   END_RUNG
   RUNG wire#w1
      R_Coil( "PB Test Air Valve" )
   END_RUNG
   RUNG wire#w1
      R_Coil( "PB Test Pneumatic 6" )
   END_RUNG
   // the same network as SCL:
   #_w1 := NOT "Machine Running" AND NOT "PB Test Mode";
   IF #_w1 AND NOT "Error" THEN
       "Flag Yellow Light" := TRUE;
       "Flag Red Light" := FALSE;
       "Flag Green Light" := FALSE;
   END_IF;
   IF #_w1 AND NOT "Error" AND NOT "Error Door Open" AND NOT "Error Door Open FC" THEN
       "Flag Kran Angin" := TRUE;
   END_IF;
   IF #_w1 THEN
       "Flag Barcode Output" := FALSE;
       "Flag Pneumatic 1" := FALSE;
       "Flag Pneumatic 2" := FALSE;
       "Flag Pneumatic 3" := FALSE;
   END_IF;
   IF #_w1 AND NOT "Section Reject" THEN
       "Flag Pneumatic 4" := FALSE;
       "Flag Pneumatic 5" := FALSE;
   END_IF;
   IF #_w1 AND NOT "Slof Manual Ready" THEN "Flag Pneumatic 6" := FALSE; END_IF;
   IF #_w1 AND NOT "Section Reject" THEN "Flag Motor" := FALSE; END_IF;
   IF #_w1 THEN
       "Flag Imaje Start" := FALSE;
       "Flag Imaje Pause" := TRUE;
       "Flag Imaje Trigger" := FALSE;
       "Flag Mesin Sebelumnya" := FALSE;
       "PB Test Pneumatic 1" := FALSE;
       "PB Test Pneumatic 2" := FALSE;
       "PB Test Pneumatic 3" := FALSE;
       "PB Test Pneumatic 4" := FALSE;
       "PB Test Pneumatic 5" := FALSE;
       "PB Test Motor" := FALSE;
       "PB Test Imaje" := FALSE;
       "PB Test Air Valve" := FALSE;
       "PB Test Pneumatic 6" := FALSE;
   END_IF;
END_REGION

REGION Network 2: Output
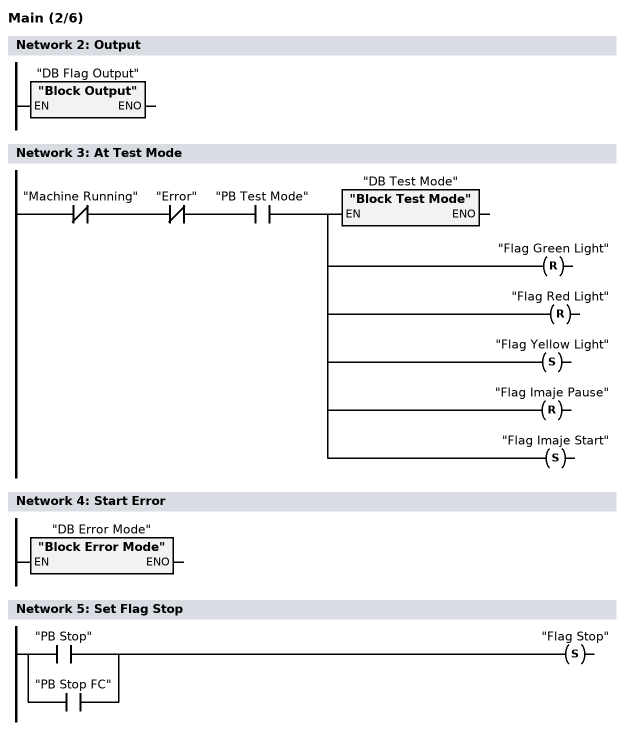
   RUNG wire#powerrail
      "DB Flag Output"()
   END_RUNG
   // the same network as SCL:
   "DB Flag Output"();   // "Block Output"
END_REGION

REGION Network 3: At Test Mode
   RUNG wire#powerrail
      I_Contact( "Machine Running" )
      I_Contact( "Error" )
      Contact( "PB Test Mode" )
      wire#w1
      "DB Test Mode"()
   END_RUNG
   RUNG wire#w1
      R_Coil( "Flag Green Light" )
   END_RUNG
   RUNG wire#w1
      R_Coil( "Flag Red Light" )
   END_RUNG
   RUNG wire#w1
      S_Coil( "Flag Yellow Light" )
   END_RUNG
   RUNG wire#w1
      R_Coil( "Flag Imaje Pause" )
   END_RUNG
   RUNG wire#w1
      S_Coil( "Flag Imaje Start" )
   END_RUNG
   // the same network as SCL:
   #_w1 := NOT "Machine Running" AND NOT "Error" AND "PB Test Mode";
   IF #_w1 THEN
       "DB Test Mode"();   // "Block Test Mode"
       "Flag Green Light" := FALSE;
       "Flag Red Light" := FALSE;
       "Flag Yellow Light" := TRUE;
       "Flag Imaje Pause" := FALSE;
       "Flag Imaje Start" := TRUE;
   END_IF;
END_REGION

REGION Network 4: Start Error
   RUNG wire#powerrail
      "DB Error Mode"()
   END_RUNG
   // the same network as SCL:
   "DB Error Mode"();   // "Block Error Mode"
END_REGION

REGION Network 5: Set Flag Stop
   RUNG wire#powerrail
      Contact( "PB Stop" )
      wire#w1
      S_Coil( "Flag Stop" )
   END_RUNG
   RUNG wire#powerrail
      Contact( "PB Stop FC" )
   END_RUNG wire#w1
   // the same network as SCL:
   IF "PB Stop" OR "PB Stop FC" THEN "Flag Stop" := TRUE; END_IF;
END_REGION

REGION Network 6: Flag Stop
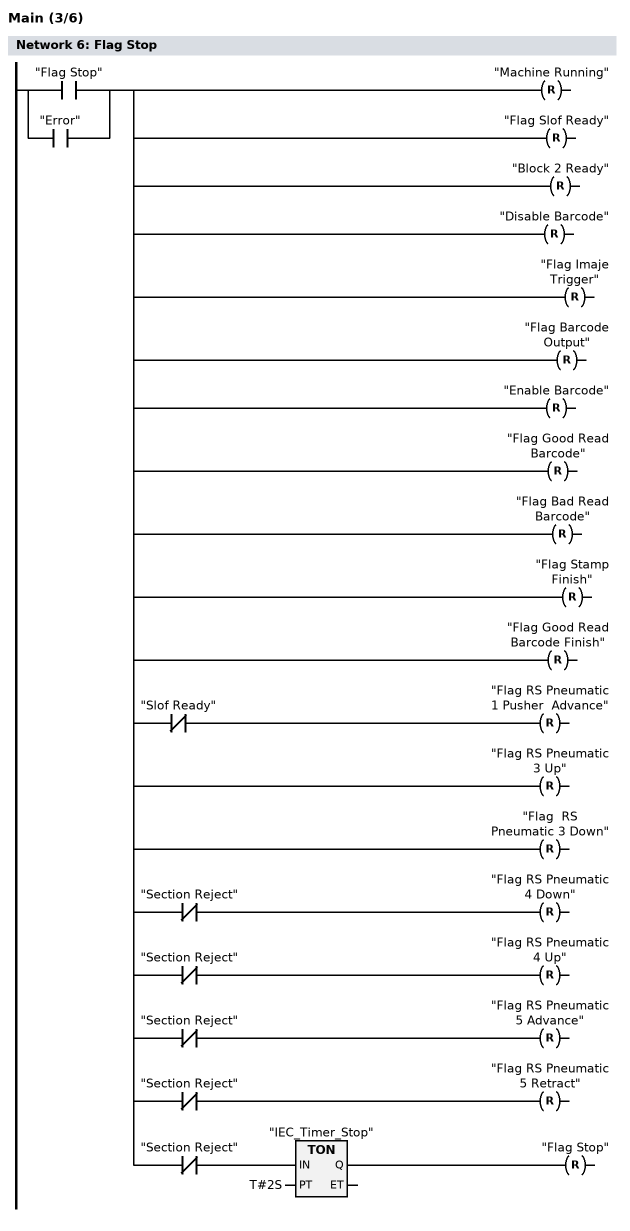
   #_w1 := "Flag Stop" OR "Error";
   IF #_w1 THEN
       "Machine Running" := FALSE;
       "Flag Slof Ready" := FALSE;
       "Block 2 Ready" := FALSE;
       "Disable Barcode" := FALSE;
       "Flag Imaje Trigger" := FALSE;
       "Flag Barcode Output" := FALSE;
       "Enable Barcode" := FALSE;
       "Flag Good Read Barcode" := FALSE;
       "Flag Bad Read Barcode" := FALSE;
       "Flag Stamp Finish" := FALSE;
       "Flag Good Read Barcode Finish" := FALSE;
   END_IF;
   IF #_w1 AND NOT "Slof Ready" THEN "Flag RS Pneumatic 1 Pusher  Advance" := FALSE; END_IF;
   IF #_w1 THEN
       "Flag RS Pneumatic 3 Up" := FALSE;
       "Flag  RS Pneumatic 3 Down" := FALSE;
   END_IF;
   IF #_w1 AND NOT "Section Reject" THEN
       "Flag RS Pneumatic 4 Down" := FALSE;
       "Flag RS Pneumatic 4 Up" := FALSE;
       "Flag RS Pneumatic 5 Advance" := FALSE;
       "Flag RS Pneumatic 5 Retract" := FALSE;
   END_IF;
   "IEC_Timer_Stop".TON(IN := #_w1 AND NOT "Section Reject", PT := T#2S);
   IF "IEC_Timer_Stop".Q THEN "Flag Stop" := FALSE; END_IF;
END_REGION

REGION Network 7: PB Run
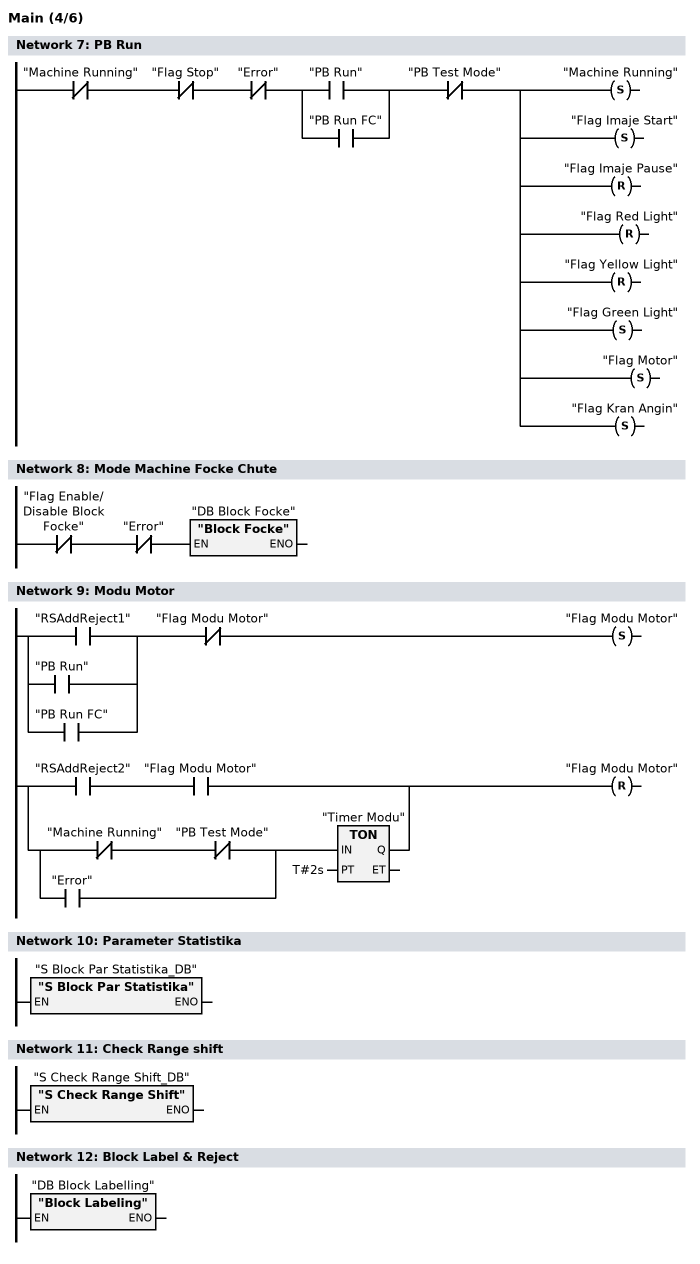
   RUNG wire#powerrail
      I_Contact( "Machine Running" )
      I_Contact( "Flag Stop" )
      I_Contact( "Error" )
      wire#w1
      Contact( "PB Run" )
      wire#w2
      I_Contact( "PB Test Mode" )
      wire#w3
      S_Coil( "Machine Running" )
   END_RUNG
   RUNG wire#w1
      Contact( "PB Run FC" )
   END_RUNG wire#w2
   RUNG wire#w3
      S_Coil( "Flag Imaje Start" )
   END_RUNG
   RUNG wire#w3
      R_Coil( "Flag Imaje Pause" )
   END_RUNG
   RUNG wire#w3
      R_Coil( "Flag Red Light" )
   END_RUNG
   RUNG wire#w3
      R_Coil( "Flag Yellow Light" )
   END_RUNG
   RUNG wire#w3
      S_Coil( "Flag Green Light" )
   END_RUNG
   RUNG wire#w3
      S_Coil( "Flag Motor" )
   END_RUNG
   RUNG wire#w3
      S_Coil( "Flag Kran Angin" )
   END_RUNG
   // the same network as SCL:
   #_w1 := NOT "Machine Running" AND NOT "Flag Stop" AND NOT "Error" AND ("PB Run" OR "PB Run FC") AND NOT "PB Test Mode";
   IF #_w1 THEN
       "Machine Running" := TRUE;
       "Flag Imaje Start" := TRUE;
       "Flag Imaje Pause" := FALSE;
       "Flag Red Light" := FALSE;
       "Flag Yellow Light" := FALSE;
       "Flag Green Light" := TRUE;
       "Flag Motor" := TRUE;
       "Flag Kran Angin" := TRUE;
   END_IF;
END_REGION

REGION Network 8: Mode Machine Focke Chute
   RUNG wire#powerrail
      I_Contact( "Flag Enable/Disable Block Focke" )
      I_Contact( "Error" )
      "DB Block Focke"()
   END_RUNG
   // the same network as SCL:
   IF NOT "Flag Enable/Disable Block Focke" AND NOT "Error" THEN
       "DB Block Focke"();   // "Block Focke"
   END_IF;
END_REGION

REGION Network 9: Modu Motor
   IF ("RSAddReject1" OR "PB Run" OR "PB Run FC") AND NOT "Flag Modu Motor" THEN
       "Flag Modu Motor" := TRUE;
   END_IF;
   "Timer Modu".TON(IN := (NOT "Machine Running" AND NOT "PB Test Mode") OR "Error", PT := T#2s);
   IF ("RSAddReject2" AND "Flag Modu Motor") OR "Timer Modu".Q THEN "Flag Modu Motor" := FALSE; END_IF;
END_REGION

REGION Network 10: Parameter Statistika
   RUNG wire#powerrail
      "S Block Par Statistika_DB"()
   END_RUNG
   // the same network as SCL:
   "S Block Par Statistika_DB"();   // "S Block Par Statistika"
END_REGION

REGION Network 11: Check Range shift
   RUNG wire#powerrail
      "S Check Range Shift_DB"()
   END_RUNG
   // the same network as SCL:
   "S Check Range Shift_DB"();   // "S Check Range Shift"
END_REGION

REGION Network 12: Block Label & Reject
   RUNG wire#powerrail
      "DB Block Labelling"()
   END_RUNG
   // the same network as SCL:
   "DB Block Labelling"();   // "Block Labeling"
END_REGION

REGION Network 13: Baca Data Statistika
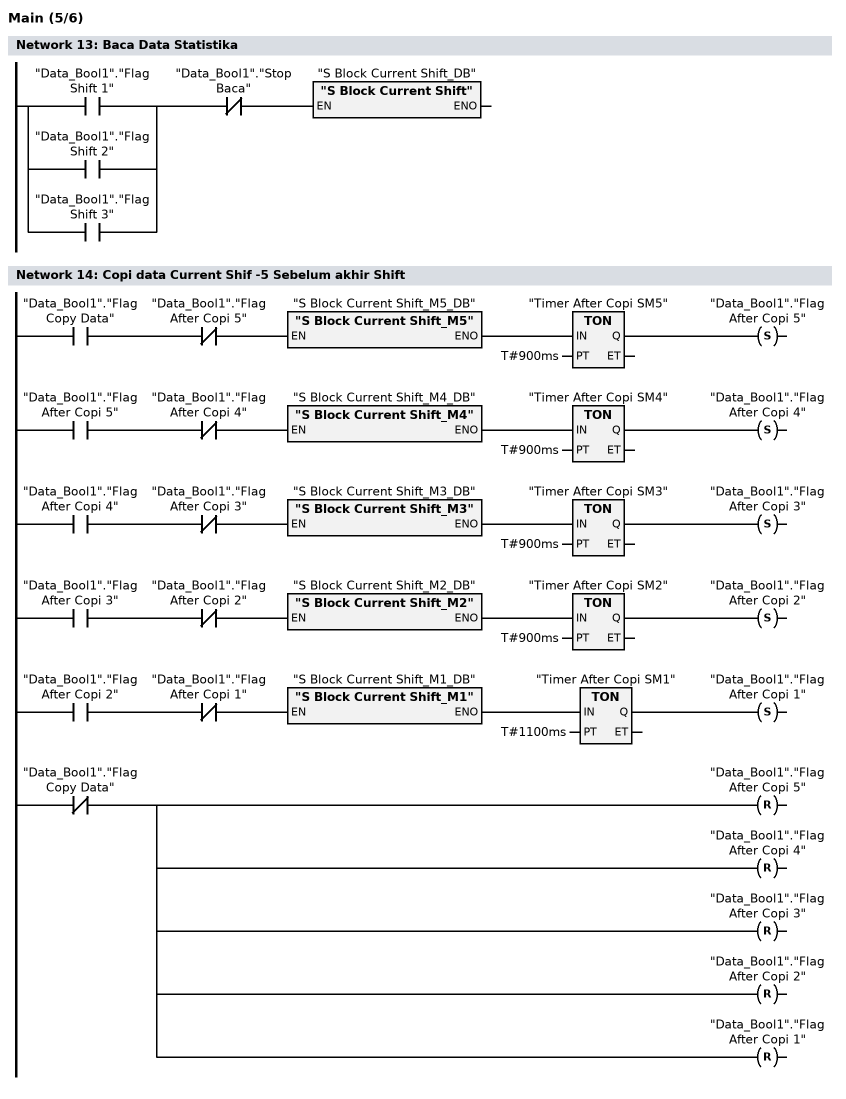
   RUNG wire#powerrail
      Contact( "Data_Bool1"."Flag Shift 1" )
      wire#w1
      I_Contact( "Data_Bool1"."Stop Baca" )
      "S Block Current Shift_DB"()
   END_RUNG
   RUNG wire#powerrail
      Contact( "Data_Bool1"."Flag Shift 2" )
   END_RUNG wire#w1
   RUNG wire#powerrail
      Contact( "Data_Bool1"."Flag Shift 3" )
   END_RUNG wire#w1
   // the same network as SCL:
   IF ("Data_Bool1"."Flag Shift 1" OR "Data_Bool1"."Flag Shift 2" OR "Data_Bool1"."Flag Shift 3") AND NOT "Data_Bool1"."Stop Baca" THEN
       "S Block Current Shift_DB"();   // "S Block Current Shift"
   END_IF;
END_REGION

REGION Network 14: Copi data Current Shif -5 Sebelum akhir Shift
   "S Block Current Shift_M5_DB"(EN := "Data_Bool1"."Flag Copy Data" AND NOT "Data_Bool1"."Flag After Copi 5",   // "S Block Current Shift_M5"
                           ENO => #_w1);
   "Timer After Copi SM5".TON(IN := #_w1, PT := T#900ms);
   IF "Timer After Copi SM5".Q THEN "Data_Bool1"."Flag After Copi 5" := TRUE; END_IF;
   "S Block Current Shift_M4_DB"(EN := "Data_Bool1"."Flag After Copi 5" AND NOT "Data_Bool1"."Flag After Copi 4",   // "S Block Current Shift_M4"
                           ENO => #_w2);
   "Timer After Copi SM4".TON(IN := #_w2, PT := T#900ms);
   IF "Timer After Copi SM4".Q THEN "Data_Bool1"."Flag After Copi 4" := TRUE; END_IF;
   "S Block Current Shift_M3_DB"(EN := "Data_Bool1"."Flag After Copi 4" AND NOT "Data_Bool1"."Flag After Copi 3",   // "S Block Current Shift_M3"
                           ENO => #_w3);
   "Timer After Copi SM3".TON(IN := #_w3, PT := T#900ms);
   IF "Timer After Copi SM3".Q THEN "Data_Bool1"."Flag After Copi 3" := TRUE; END_IF;
   "S Block Current Shift_M2_DB"(EN := "Data_Bool1"."Flag After Copi 3" AND NOT "Data_Bool1"."Flag After Copi 2",   // "S Block Current Shift_M2"
                           ENO => #_w4);
   "Timer After Copi SM2".TON(IN := #_w4, PT := T#900ms);
   IF "Timer After Copi SM2".Q THEN "Data_Bool1"."Flag After Copi 2" := TRUE; END_IF;
   "S Block Current Shift_M1_DB"(EN := "Data_Bool1"."Flag After Copi 2" AND NOT "Data_Bool1"."Flag After Copi 1",   // "S Block Current Shift_M1"
                           ENO => #_w5);
   "Timer After Copi SM1".TON(IN := #_w5, PT := T#1100ms);
   IF "Timer After Copi SM1".Q THEN "Data_Bool1"."Flag After Copi 1" := TRUE; END_IF;
   IF NOT "Data_Bool1"."Flag Copy Data" THEN
       "Data_Bool1"."Flag After Copi 5" := FALSE;
       "Data_Bool1"."Flag After Copi 4" := FALSE;
       "Data_Bool1"."Flag After Copi 3" := FALSE;
       "Data_Bool1"."Flag After Copi 2" := FALSE;
       "Data_Bool1"."Flag After Copi 1" := FALSE;
   END_IF;
END_REGION

REGION Network 15: Hapus Data Current shift
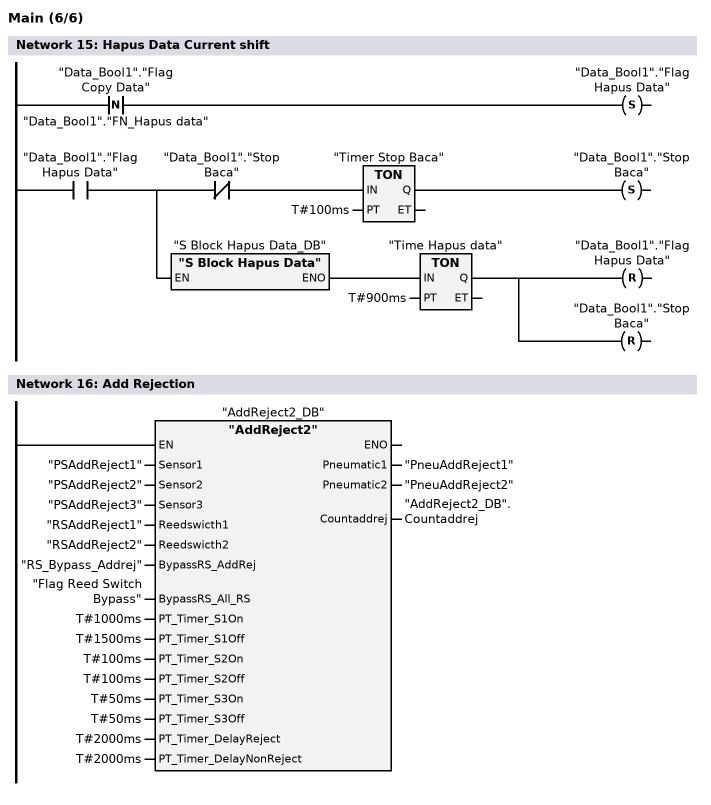
   #_w1 := NOT "Data_Bool1"."Flag Copy Data" AND "Data_Bool1"."FN_Hapus data";   // falling edge of "Data_Bool1"."Flag Copy Data"
   "Data_Bool1"."FN_Hapus data" := "Data_Bool1"."Flag Copy Data";
   IF #_w1 THEN "Data_Bool1"."Flag Hapus Data" := TRUE; END_IF;
   "Timer Stop Baca".TON(IN := "Data_Bool1"."Flag Hapus Data" AND NOT "Data_Bool1"."Stop Baca", PT := T#100ms);
   IF "Timer Stop Baca".Q THEN "Data_Bool1"."Stop Baca" := TRUE; END_IF;
   "S Block Hapus Data_DB"(EN := "Data_Bool1"."Flag Hapus Data", ENO => #_w2);   // "S Block Hapus Data"
   "Time Hapus data".TON(IN := #_w2, PT := T#900ms);
   IF "Time Hapus data".Q THEN
       "Data_Bool1"."Flag Hapus Data" := FALSE;
       "Data_Bool1"."Stop Baca" := FALSE;
   END_IF;
END_REGION

REGION Network 16: Add Rejection
   RUNG wire#powerrail
      "AddReject2_DB"(Sensor1 := "PSAddReject1", Sensor2 := "PSAddReject2", Sensor3 := "PSAddReject3", Reedswicth1 := "RSAddReject1", Reedswicth2 := "RSAddReject2", BypassRS_AddRej := "RS_Bypass_Addrej", BypassRS_All_RS := "Flag Reed Switch Bypass", PT_Timer_S1On := T#1000ms, PT_Timer_S1Off := T#1500ms, PT_Timer_S2On := T#100ms, PT_Timer_S2Off := T#100ms, PT_Timer_S3On := T#50ms, PT_Timer_S3Off := T#50ms, PT_Timer_DelayReject := T#2000ms, PT_Timer_DelayNonReject := T#2000ms, Pneumatic1 => "PneuAddReject1", Pneumatic2 => "PneuAddReject2", Countaddrej => "AddReject2_DB".Countaddrej)
   END_RUNG
   // the same network as SCL:
   "AddReject2_DB"(Sensor1 := "PSAddReject1",   // "AddReject2"
                   Sensor2 := "PSAddReject2",
                   Sensor3 := "PSAddReject3",
                   Reedswicth1 := "RSAddReject1",
                   Reedswicth2 := "RSAddReject2",
                   BypassRS_AddRej := "RS_Bypass_Addrej",
                   BypassRS_All_RS := "Flag Reed Switch Bypass",
                   PT_Timer_S1On := T#1000ms,
                   PT_Timer_S1Off := T#1500ms,
                   PT_Timer_S2On := T#100ms,
                   PT_Timer_S2Off := T#100ms,
                   PT_Timer_S3On := T#50ms,
                   PT_Timer_S3Off := T#50ms,
                   PT_Timer_DelayReject := T#2000ms,
                   PT_Timer_DelayNonReject := T#2000ms,
                   Pneumatic1 => "PneuAddReject1",
                   Pneumatic2 => "PneuAddReject2",
                   Countaddrej => "AddReject2_DB".Countaddrej);
END_REGION
END_ORGANIZATION_BLOCK

(* ===== HMI "HMI_RT_1" =====
system functions are stored by id; their names below are inferred from use
connection "HMI_connection": ETHERNET, SMART_S7_1200_OMS

HMI tags "Default tag table"
   "Tag_ScreenNumber" : UInt, internal
      on ChangeValue: ActivateScreenByNumber("Tag_ScreenNumber", 0)
   "PB Test Pneumatic 1" : Bool = PLC "PB Test Pneumatic 1" AT %M205.1, 1 s
   "PB Test Pneumatic 2" : Bool = PLC "PB Test Pneumatic 2" AT %M205.2, 1 s
   "PB Test Pneumatic 3" : Bool = PLC "PB Test Pneumatic 3" AT %M205.3, 1 s
   "PB Test Pneumatic 4" : Bool = PLC "PB Test Pneumatic 4" AT %M205.4, 1 s
   "PB Test Pneumatic 5" : Bool = PLC "PB Test Pneumatic 5" AT %M205.5, 1 s
   "PB Test Motor" : Bool = PLC "PB Test Motor" AT %M205.7, 1 s
   "PB Test Manual Servo" : Bool = PLC "PB Test Manual Servo" AT %M205.6, 1 s
   "Machine Running" : Bool = PLC "Machine Running" AT %M200.0, 1 s
   "Flag Imaje Start" : Bool = PLC "Flag Imaje Start" AT %M212.0, 1 s
   "Reset Counter" : Bool = PLC "Reset Counter" AT %M200.1, 1 s
   "PB Test Mode" : Bool = PLC "PB Test Mode" AT %M205.0, 1 s
   "Flag Ejector Jalan" : Bool = PLC "Flag Ejector Jalan" AT %M230.3, 1 s
   "Error Group" : Word = PLC "Error Group" AT %MW4, 1 s
   "PB Test Imaje" : Bool = PLC "PB Test Imaje" AT %M206.0, 1 s
   "PB Test Air Valve" : Bool = PLC "PB Test Air Valve" AT %M206.1, 1 s
   "Flag Barcode HMI" : Bool = PLC "Flag Enable/Disable Barcode HMI" AT %M30.0, 1 s
   "Flag Enable/Disable Error Chute 3 Way" : Bool = PLC "Flag Enable/Disable Error Chute 3 Way" AT %M30.1, 1 s
   "Flag Parameter Page" : Bool = PLC "Flag Parameter Page" AT %M232.6, 1 s
   "Flag Main Page" : Bool = PLC "Flag Main Page" AT %M232.7, 1 s
   "HMI_Tag_1" : Word AT %DB39.DBW0, 1 s
   "HMI_Error_Cont" : Word AT %DB40.DBW0, 1 s
   "Flag Teach In Barcode" : Bool = PLC "Flag Teach In Barcode" AT %M212.4, 1 s
   "Teach In Barcode" : Bool = PLC "Teach In Barcode" AT %Q0.5, 1 s
   "Flag Heater Error HMI" : Bool = PLC "Flag Heater Error HMI" AT %M30.2, 1 s
   "Flag Pneumatic Bypass" : Bool = PLC "Flag Reed Switch Bypass" AT %M30.3, 1 s
   "Flag Enable/Disable Error Door Open" : Bool = PLC "Flag Enable/Disable Error Door Open" AT %M30.5, 1 s
   "Flag Enable/Disable Block Focke" : Bool = PLC "Flag Enable/Disable Block Focke" AT %M30.6, 1 s
   "Flag Enable/Disable Error Chute Before Heating Roll" : Bool = PLC "Flag Enable/Disable Error Chute Before Heating Roll" AT %M30.4, 1 s
   "Flag Machine Bypass" : Bool = PLC "Flag Machine Bypass" AT %M30.7, 1 s
   "RS Bypass Pneumatic 1" : Bool = PLC "RS Bypass Pneumatic 1" AT %M31.0, 1 s
   "RS Bypass Pneumatic 3" : Bool = PLC "RS Bypass Pneumatic 3" AT %M31.1, 1 s
   "RS Bypass Pneumatic 4" : Bool = PLC "RS Bypass Pneumatic 4" AT %M31.2, 1 s
   "RS Bypass Pneumatic 5" : Bool = PLC "RS Bypass Pneumatic 5" AT %M31.3, 1 s
   "PB Test Pneumatic 6" : Bool = PLC "PB Test Pneumatic 6" AT %M206.2, 1 s
   "PB Test Conveyor" : Bool = PLC "PB Test Conveyor" AT %M206.3, 1 s
   "Flag Enable/Disable Flow to Reject" : Bool = PLC "Flag Enable/Disable Flow to Reject" AT %M31.5, 1 s
   "PB Test Motor Coveyor Pusher" : Bool = PLC "PB Test Motor Coveyor Pusher" AT %M206.4, 1 s
   "PB Test Motor Heating Roll" : Bool = PLC "PB Test Motor Heating Roll" AT %M206.5, 1 s
   "Flag Enable/Disable Heating Roll" : Bool = PLC "Flag Enable/Disable Heating Roll" AT %M31.6, 1 s
   "Flag Enable/Disable Reject Outfeed" : Bool = PLC "Flag Enable/Disable Reject Outfeed" AT %M31.7, 1 s
   "Data_DTL1_Output" : DTL = PLC Data_DTL1.Output, 1 s
   "Data_DTL1_Cur_ShiftA" : DTL = PLC Data_DTL1.Cur_ShiftA, 1 s
   "Data_DTL1_Cur_ShiftB" : DTL = PLC Data_DTL1.Cur_ShiftB, 1 s
   "Data_IntData_Input Sloft" : UDInt = PLC Data_IntData."Input Sloft", 1 s
   "Data_IntData_Tot Out Slof" : UDInt = PLC Data_IntData."Tot Out Slof", 1 s
   "Data_IntData_Good R" : UDInt = PLC Data_IntData."Good R", 1 s
   "Data_IntData_Reject Out S" : UDInt = PLC Data_IntData."Reject Out S", 1 s
   "Data_IntData_Bad R" : UDInt = PLC Data_IntData."Bad R", 1 s
   "Data_Real_% Total Output[0]" : Real = PLC Data_Real."% Total Output"[0], 1 s
   "Data_Real_%Good Read[0]" : Real = PLC Data_Real."%Good Read"[0], 1 s
   "Data_Real_% Reject Out Stop[0]" : Real = PLC Data_Real."% Reject Out Stop"[0], 1 s
   "Data_Real_%Bad Read[0]" : Real = PLC Data_Real."%Bad Read"[0], 1 s
   "Data_DTL1_Cur_ShiftA_1" : DTL = PLC Data_DTL1.Cur_ShiftA_1, 1 s
   "Data_DTL1_Cur_ShiftB_1" : DTL = PLC Data_DTL1.Cur_ShiftB_1, 1 s
   "Data_DTL1_Cur_ShiftA_2" : DTL = PLC Data_DTL1.Cur_ShiftA_2, 1 s
   "Data_DTL1_Cur_ShiftB_2" : DTL = PLC Data_DTL1.Cur_ShiftB_2, 1 s
   "Data_DTL1_Cur_ShiftA_3" : DTL = PLC Data_DTL1.Cur_ShiftA_3, 1 s
   "Data_DTL1_Cur_ShiftB_3" : DTL = PLC Data_DTL1.Cur_ShiftB_3, 1 s
   "Data_DTL1_Cur_ShiftA_4" : DTL = PLC Data_DTL1.Cur_ShiftA_4, 1 s
   "Data_DTL1_Cur_ShiftB_4" : DTL = PLC Data_DTL1.Cur_ShiftB_4, 1 s
   "Data_IntData_Input Sloft_1" : UDInt = PLC Data_IntData."Input Sloft_1", 1 s
   "Data_IntData_Tot Out Slof_1" : UDInt = PLC Data_IntData."Tot Out Slof_1", 1 s
   "Data_IntData_Good R_1" : UDInt = PLC Data_IntData."Good R_1", 1 s
   "Data_IntData_Reject Out S_1" : UDInt = PLC Data_IntData."Reject Out S_1", 1 s
   "Data_IntData_Bad R_1" : UDInt = PLC Data_IntData."Bad R_1", 1 s
   "Data_Real_% Total Output[1]" : Real = PLC Data_Real."% Total Output"[1], 1 s
   "Data_Real_%Good Read[1]" : Real = PLC Data_Real."%Good Read"[1], 1 s
   "Data_Real_% Reject Out Stop[1]" : Real = PLC Data_Real."% Reject Out Stop"[1], 1 s
   "Data_Real_%Bad Read[1]" : Real = PLC Data_Real."%Bad Read"[1], 1 s
   "Data_Real_% Total Output[2]" : Real = PLC Data_Real."% Total Output"[2], 1 s
   "Data_Real_%Good Read[2]" : Real = PLC Data_Real."%Good Read"[2], 1 s
   "Data_Real_% Reject Out Stop[2]" : Real = PLC Data_Real."% Reject Out Stop"[2], 1 s
   "Data_Real_%Bad Read[2]" : Real = PLC Data_Real."%Bad Read"[2], 1 s
   "Data_IntData_Input Sloft_2" : UDInt = PLC Data_IntData."Input Sloft_2", 1 s
   "Data_IntData_Tot Out Slof_2" : UDInt = PLC Data_IntData."Tot Out Slof_2", 1 s
   "Data_IntData_Good R_2" : UDInt = PLC Data_IntData."Good R_2", 1 s
   "Data_IntData_Reject Out S_2" : UDInt = PLC Data_IntData."Reject Out S_2", 1 s
   "Data_IntData_Bad R_2" : UDInt = PLC Data_IntData."Bad R_2", 1 s
   "Data_IntData_Input Sloft_3" : UDInt = PLC Data_IntData."Input Sloft_3", 1 s
   "Data_IntData_Tot Out Slof_3" : UDInt = PLC Data_IntData."Tot Out Slof_3", 1 s
   "Data_IntData_Good R_3" : UDInt = PLC Data_IntData."Good R_3", 1 s
   "Data_IntData_Reject Out S_3" : UDInt = PLC Data_IntData."Reject Out S_3", 1 s
   "Data_IntData_Bad R_3" : UDInt = PLC Data_IntData."Bad R_3", 1 s
   "Data_Real_% Total Output[3]" : Real = PLC Data_Real."% Total Output"[3], 1 s
   "Data_Real_%Good Read[3]" : Real = PLC Data_Real."%Good Read"[3], 1 s
   "Data_Real_% Reject Out Stop[3]" : Real = PLC Data_Real."% Reject Out Stop"[3], 1 s
   "Data_Real_%Bad Read[3]" : Real = PLC Data_Real."%Bad Read"[3], 1 s
   "Data_Real_% Total Output[4]" : Real = PLC Data_Real."% Total Output"[4], 1 s
   "Data_Real_%Good Read[4]" : Real = PLC Data_Real."%Good Read"[4], 1 s
   "Data_Real_% Reject Out Stop[4]" : Real = PLC Data_Real."% Reject Out Stop"[4], 1 s
   "Data_Real_%Bad Read[4]" : Real = PLC Data_Real."%Bad Read"[4], 1 s
   "Data_IntData_Input Sloft_4" : UDInt = PLC Data_IntData."Input Sloft_4", 1 s
   "Data_IntData_Tot Out Slof_4" : UDInt = PLC Data_IntData."Tot Out Slof_4", 1 s
   "Data_IntData_Good R_4" : UDInt = PLC Data_IntData."Good R_4", 1 s
   "Data_IntData_Reject Out S_4" : UDInt = PLC Data_IntData."Reject Out S_4", 1 s
   "Data_IntData_Bad R_4" : UDInt = PLC Data_IntData."Bad R_4", 1 s
   "Data_IntData_Input Sloft_5" : UDInt = PLC Data_IntData."Input Sloft_5", 1 s
   "Data_IntData_Tot Out Slof_5" : UDInt = PLC Data_IntData."Tot Out Slof_5", 1 s
   "Data_IntData_Good R_5" : UDInt = PLC Data_IntData."Good R_5", 1 s
   "Data_IntData_Reject Out S_5" : UDInt = PLC Data_IntData."Reject Out S_5", 1 s
   "Data_IntData_Bad R_5" : UDInt = PLC Data_IntData."Bad R_5", 1 s
   "Data_Real_% Total Output[5]" : Real = PLC Data_Real."% Total Output"[5], 1 s
   "Data_Real_%Good Read[5]" : Real = PLC Data_Real."%Good Read"[5], 1 s
   "Data_Real_% Reject Out Stop[5]" : Real = PLC Data_Real."% Reject Out Stop"[5], 1 s
   "Data_Real_%Bad Read[5]" : Real = PLC Data_Real."%Bad Read"[5], 1 s
   "Data_DTLData_DTL_Imaje Er.HOUR" : USInt = PLC Data_DTLData."DTL_Imaje Er".HOUR, 1 s
   "Data_DTLData_DTL_Imaje Er.MINUTE" : USInt = PLC Data_DTLData."DTL_Imaje Er".MINUTE, 1 s
   "Data_DTLData_DTL_Imaje Er.SECOND" : USInt = PLC Data_DTLData."DTL_Imaje Er".SECOND, 1 s
   "Data_DTLData_DTL_Imaje Not In Position[0].HOUR" : USInt = PLC Data_DTLData."DTL_Imaje Not In Position"[0].HOUR, 1 s
   "Data_DTLData_DTL_Paper R Out[0].HOUR" : USInt = PLC Data_DTLData."DTL_Paper R Out"[0].HOUR, 1 s
   "Data_DTLData_DTL_Paper R Out[0].MINUTE" : USInt = PLC Data_DTLData."DTL_Paper R Out"[0].MINUTE, 1 s
   "Data_DTLData_DTL_Paper R Out[0].SECOND" : USInt = PLC Data_DTLData."DTL_Paper R Out"[0].SECOND, 1 s
   "Data_DTLData_DTL_Imaje Not In Position[0].MINUTE" : USInt = PLC Data_DTLData."DTL_Imaje Not In Position"[0].MINUTE, 1 s
   "Data_DTLData_DTL_Imaje Not In Position[0].SECOND" : USInt = PLC Data_DTLData."DTL_Imaje Not In Position"[0].SECOND, 1 s
   "Data_DTLData_DTL_Sloft Jam1.HOUR" : USInt = PLC Data_DTLData."DTL_Sloft Jam1".HOUR, 1 s
   "Data_DTLData_DTL_Sloft Jam1.MINUTE" : USInt = PLC Data_DTLData."DTL_Sloft Jam1".MINUTE, 1 s
   "Data_DTLData_DTL_Sloft Jam1.SECOND" : USInt = PLC Data_DTLData."DTL_Sloft Jam1".SECOND, 1 s
   "Data_DTLData_DTL_Down Stop.HOUR" : USInt = PLC Data_DTLData."DTL_Down Stop".HOUR, 1 s
   "Data_DTLData_DTL_Down Stop.MINUTE" : USInt = PLC Data_DTLData."DTL_Down Stop".MINUTE, 1 s
   "Data_DTLData_DTL_Down Stop.SECOND" : USInt = PLC Data_DTLData."DTL_Down Stop".SECOND, 1 s
   "Data_DTLData_DTL_RS Pneu Er.HOUR" : USInt = PLC Data_DTLData."DTL_RS Pneu Er".HOUR, 1 s
   "Data_DTLData_DTL_RS Pneu Er.MINUTE" : USInt = PLC Data_DTLData."DTL_RS Pneu Er".MINUTE, 1 s
   "Data_DTLData_DTL_RS Pneu Er.SECOND" : USInt = PLC Data_DTLData."DTL_RS Pneu Er".SECOND, 1 s
   "Data_DTLData_DTL_Imaje Er_1.HOUR" : USInt = PLC Data_DTLData."DTL_Imaje Er_1".HOUR, 1 s
   "Data_DTLData_DTL_Imaje Er_1.MINUTE" : USInt = PLC Data_DTLData."DTL_Imaje Er_1".MINUTE, 1 s
   "Data_DTLData_DTL_Imaje Er_1.SECOND" : USInt = PLC Data_DTLData."DTL_Imaje Er_1".SECOND, 1 s
   "Data_DTLData_DTL_Paper R Out[1].HOUR" : USInt = PLC Data_DTLData."DTL_Paper R Out"[1].HOUR, 1 s
   "Data_DTLData_DTL_Imaje Not In Position[1].MINUTE" : USInt = PLC Data_DTLData."DTL_Imaje Not In Position"[1].MINUTE, 1 s
   "Data_DTLData_DTL_Paper R Out[1].SECOND" : USInt = PLC Data_DTLData."DTL_Paper R Out"[1].SECOND, 1 s
   "Data_DTLData_DTL_Paper R Out[1].MINUTE" : USInt = PLC Data_DTLData."DTL_Paper R Out"[1].MINUTE, 1 s
   "Data_DTLData_DTL_Imaje Not In Position[2].HOUR" : USInt = PLC Data_DTLData."DTL_Imaje Not In Position"[2].HOUR, 1 s
   "Data_DTLData_DTL_Sloft Jam1_1.HOUR" : USInt = PLC Data_DTLData."DTL_Sloft Jam1_1".HOUR, 1 s
   "Data_DTLData_DTL_Sloft Jam1_1.MINUTE" : USInt = PLC Data_DTLData."DTL_Sloft Jam1_1".MINUTE, 1 s
   "Data_DTLData_DTL_Sloft Jam1_1.SECOND" : USInt = PLC Data_DTLData."DTL_Sloft Jam1_1".SECOND, 1 s
   "Data_DTLData_DTL_Down Stop_1.HOUR" : USInt = PLC Data_DTLData."DTL_Down Stop_1".HOUR, 1 s
   "Data_DTLData_DTL_Down Stop_1.MINUTE" : USInt = PLC Data_DTLData."DTL_Down Stop_1".MINUTE, 1 s
   "Data_DTLData_DTL_Down Stop_1.SECOND" : USInt = PLC Data_DTLData."DTL_Down Stop_1".SECOND, 1 s
   "Data_DTLData_DTL_RS Pneu Er_1.HOUR" : USInt = PLC Data_DTLData."DTL_RS Pneu Er_1".HOUR, 1 s
   "Data_DTLData_DTL_RS Pneu Er_1.MINUTE" : USInt = PLC Data_DTLData."DTL_RS Pneu Er_1".MINUTE, 1 s
   "Data_DTLData_DTL_RS Pneu Er_1.SECOND" : USInt = PLC Data_DTLData."DTL_RS Pneu Er_1".SECOND, 1 s
   "Data_DTLData_DTL_Imaje Er_2.HOUR" : USInt = PLC Data_DTLData."DTL_Imaje Er_2".HOUR, 1 s
   "Data_DTLData_DTL_Imaje Er_2.MINUTE" : USInt = PLC Data_DTLData."DTL_Imaje Er_2".MINUTE, 1 s
   "Data_DTLData_DTL_Imaje Er_2.SECOND" : USInt = PLC Data_DTLData."DTL_Imaje Er_2".SECOND, 1 s
   "Data_DTLData_DTL_Paper R Out[2].HOUR" : USInt = PLC Data_DTLData."DTL_Paper R Out"[2].HOUR, 1 s
   "Data_DTLData_DTL_Paper R Out[2].MINUTE" : USInt = PLC Data_DTLData."DTL_Paper R Out"[2].MINUTE, 1 s
   "Data_DTLData_DTL_Paper R Out[2].SECOND" : USInt = PLC Data_DTLData."DTL_Paper R Out"[2].SECOND, 1 s
   "Data_DTLData_DTL_Imaje Not In Position[2].MINUTE" : USInt = PLC Data_DTLData."DTL_Imaje Not In Position"[2].MINUTE, 1 s
   "Data_DTLData_DTL_Imaje Not In Position[2].SECOND" : USInt = PLC Data_DTLData."DTL_Imaje Not In Position"[2].SECOND, 1 s
   "Data_DTLData_DTL_Sloft Jam1_3.HOUR" : USInt = PLC Data_DTLData."DTL_Sloft Jam1_3".HOUR, 1 s
   "Data_DTLData_DTL_Sloft Jam1_3.MINUTE" : USInt = PLC Data_DTLData."DTL_Sloft Jam1_3".MINUTE, 1 s
   "Data_DTLData_DTL_Sloft Jam1_3.SECOND" : USInt = PLC Data_DTLData."DTL_Sloft Jam1_3".SECOND, 1 s
   "Data_DTLData_DTL_Down Stop_3.HOUR" : USInt = PLC Data_DTLData."DTL_Down Stop_3".HOUR, 1 s
   "Data_DTLData_DTL_Down Stop_3.MINUTE" : USInt = PLC Data_DTLData."DTL_Down Stop_3".MINUTE, 1 s
   "Data_DTLData_DTL_Down Stop_3.SECOND" : USInt = PLC Data_DTLData."DTL_Down Stop_3".SECOND, 1 s
   "Data_DTLData_DTL_RS Pneu Er_3.HOUR" : USInt = PLC Data_DTLData."DTL_RS Pneu Er_3".HOUR, 1 s
   "Data_DTLData_DTL_Imaje Not In Position[1].HOUR" : USInt = PLC Data_DTLData."DTL_Imaje Not In Position"[1].HOUR, 1 s
   "Data_DTLData_DTL_Imaje Not In Position[1].SECOND" : USInt = PLC Data_DTLData."DTL_Imaje Not In Position"[1].SECOND, 1 s
   "Data_DTLData_DTL_RS Pneu Er_3.MINUTE" : USInt = PLC Data_DTLData."DTL_RS Pneu Er_3".MINUTE, 1 s
   "Data_DTLData_DTL_RS Pneu Er_3.SECOND" : USInt = PLC Data_DTLData."DTL_RS Pneu Er_3".SECOND, 1 s
   "Data_DTLData_DTL_Sloft Jam1_2.HOUR" : USInt = PLC Data_DTLData."DTL_Sloft Jam1_2".HOUR, 1 s
   "Data_DTLData_DTL_Sloft Jam1_2.MINUTE" : USInt = PLC Data_DTLData."DTL_Sloft Jam1_2".MINUTE, 1 s
   "Data_DTLData_DTL_Sloft Jam1_2.SECOND" : USInt = PLC Data_DTLData."DTL_Sloft Jam1_2".SECOND, 1 s
   "Data_DTLData_DTL_Down Stop_2.HOUR" : USInt = PLC Data_DTLData."DTL_Down Stop_2".HOUR, 1 s
   "Data_DTLData_DTL_Down Stop_2.MINUTE" : USInt = PLC Data_DTLData."DTL_Down Stop_2".MINUTE, 1 s
   "Data_DTLData_DTL_Down Stop_2.SECOND" : USInt = PLC Data_DTLData."DTL_Down Stop_2".SECOND, 1 s
   "Data_DTLData_DTL_RS Pneu Er_2.HOUR" : USInt = PLC Data_DTLData."DTL_RS Pneu Er_2".HOUR, 1 s
   "Data_DTLData_DTL_RS Pneu Er_2.MINUTE" : USInt = PLC Data_DTLData."DTL_RS Pneu Er_2".MINUTE, 1 s
   "Data_DTLData_DTL_RS Pneu Er_2.SECOND" : USInt = PLC Data_DTLData."DTL_RS Pneu Er_2".SECOND, 1 s
   "Data_DTL1_Cur_ShiftA_5" : DTL = PLC Data_DTL1.Cur_ShiftA_5, 1 s
   "Data_DTL1_Cur_ShiftB_5" : DTL = PLC Data_DTL1.Cur_ShiftB_5, 1 s
   "Data_DTLData_DTL_Imaje Er_5.HOUR" : USInt = PLC Data_DTLData."DTL_Imaje Er_5".HOUR, 1 s
   "Data_DTLData_DTL_Imaje Er_5.MINUTE" : USInt = PLC Data_DTLData."DTL_Imaje Er_5".MINUTE, 1 s
   "Data_DTLData_DTL_Imaje Er_5.SECOND" : USInt = PLC Data_DTLData."DTL_Imaje Er_5".SECOND, 1 s
   "Data_DTLData_DTL_Paper R Out[5].HOUR" : USInt = PLC Data_DTLData."DTL_Paper R Out"[5].HOUR, 1 s
   "Data_DTLData_DTL_Paper R Out[5].MINUTE" : USInt = PLC Data_DTLData."DTL_Paper R Out"[5].MINUTE, 1 s
   "Data_DTLData_DTL_Paper R Out[5].SECOND" : USInt = PLC Data_DTLData."DTL_Paper R Out"[5].SECOND, 1 s
   "Data_DTLData_DTL_Imaje Not In Position[5].HOUR" : USInt = PLC Data_DTLData."DTL_Imaje Not In Position"[5].HOUR, 1 s
   "Data_DTLData_DTL_Imaje Not In Position[5].MINUTE" : USInt = PLC Data_DTLData."DTL_Imaje Not In Position"[5].MINUTE, 1 s
   "Data_DTLData_DTL_Imaje Not In Position[5].SECOND" : USInt = PLC Data_DTLData."DTL_Imaje Not In Position"[5].SECOND, 1 s
   "Data_DTLData_DTL_Sloft Jam1_5.HOUR" : USInt = PLC Data_DTLData."DTL_Sloft Jam1_5".HOUR, 1 s
   "Data_DTLData_DTL_Sloft Jam1_5.MINUTE" : USInt = PLC Data_DTLData."DTL_Sloft Jam1_5".MINUTE, 1 s
   "Data_DTLData_DTL_Sloft Jam1_5.SECOND" : USInt = PLC Data_DTLData."DTL_Sloft Jam1_5".SECOND, 1 s
   "Data_DTLData_DTL_Down Stop_5.HOUR" : USInt = PLC Data_DTLData."DTL_Down Stop_5".HOUR, 1 s
   "Data_DTLData_DTL_Down Stop_5.MINUTE" : USInt = PLC Data_DTLData."DTL_Down Stop_5".MINUTE, 1 s
   "Data_DTLData_DTL_Down Stop_5.SECOND" : USInt = PLC Data_DTLData."DTL_Down Stop_5".SECOND, 1 s
   "Data_DTLData_DTL_RS Pneu Er_5.HOUR" : USInt = PLC Data_DTLData."DTL_RS Pneu Er_5".HOUR, 1 s
   "Data_DTLData_DTL_RS Pneu Er_5.MINUTE" : USInt = PLC Data_DTLData."DTL_RS Pneu Er_5".MINUTE, 1 s
   "Data_DTLData_DTL_RS Pneu Er_5.SECOND" : USInt = PLC Data_DTLData."DTL_RS Pneu Er_5".SECOND, 1 s
   "Data_DTLData_DTL_Imaje Er_4.HOUR" : USInt = PLC Data_DTLData."DTL_Imaje Er_4".HOUR, 1 s
   "Data_DTLData_DTL_Imaje Er_4.MINUTE" : USInt = PLC Data_DTLData."DTL_Imaje Er_4".MINUTE, 1 s
   "Data_DTLData_DTL_Imaje Er_4.SECOND" : USInt = PLC Data_DTLData."DTL_Imaje Er_4".SECOND, 1 s
   "Data_DTLData_DTL_Paper R Out[4].HOUR" : USInt = PLC Data_DTLData."DTL_Paper R Out"[4].HOUR, 1 s
   "Data_DTLData_DTL_Paper R Out[4].MINUTE" : USInt = PLC Data_DTLData."DTL_Paper R Out"[4].MINUTE, 1 s
   "Data_DTLData_DTL_Paper R Out[4].SECOND" : USInt = PLC Data_DTLData."DTL_Paper R Out"[4].SECOND, 1 s
   "Data_DTLData_DTL_Imaje Not In Position[4].HOUR" : USInt = PLC Data_DTLData."DTL_Imaje Not In Position"[4].HOUR, 1 s
   "Data_DTLData_DTL_Imaje Not In Position[4].MINUTE" : USInt = PLC Data_DTLData."DTL_Imaje Not In Position"[4].MINUTE, 1 s
   "Data_DTLData_DTL_Imaje Not In Position[4].SECOND" : USInt = PLC Data_DTLData."DTL_Imaje Not In Position"[4].SECOND, 1 s
   "Data_DTLData_DTL_Sloft Jam1_4.HOUR" : USInt = PLC Data_DTLData."DTL_Sloft Jam1_4".HOUR, 1 s
   "Data_DTLData_DTL_Sloft Jam1_4.MINUTE" : USInt = PLC Data_DTLData."DTL_Sloft Jam1_4".MINUTE, 1 s
   "Data_DTLData_DTL_Sloft Jam1_4.SECOND" : USInt = PLC Data_DTLData."DTL_Sloft Jam1_4".SECOND, 1 s
   "Data_DTLData_DTL_Down Stop_4.HOUR" : USInt = PLC Data_DTLData."DTL_Down Stop_4".HOUR, 1 s
   "Data_DTLData_DTL_Down Stop_4.MINUTE" : USInt = PLC Data_DTLData."DTL_Down Stop_4".MINUTE, 1 s
   "Data_DTLData_DTL_Down Stop_4.SECOND" : USInt = PLC Data_DTLData."DTL_Down Stop_4".SECOND, 1 s
   "Data_DTLData_DTL_RS Pneu Er_4.HOUR" : USInt = PLC Data_DTLData."DTL_RS Pneu Er_4".HOUR, 1 s
   "Data_DTLData_DTL_RS Pneu Er_4.MINUTE" : USInt = PLC Data_DTLData."DTL_RS Pneu Er_4".MINUTE, 1 s
   "Data_DTLData_DTL_RS Pneu Er_4.SECOND" : USInt = PLC Data_DTLData."DTL_RS Pneu Er_4".SECOND, 1 s
   "Data_DTLData_DTL_Imaje Er_3.HOUR" : USInt = PLC Data_DTLData."DTL_Imaje Er_3".HOUR, 1 s
   "Data_DTLData_DTL_Imaje Er_3.MINUTE" : USInt = PLC Data_DTLData."DTL_Imaje Er_3".MINUTE, 1 s
   "Data_DTLData_DTL_Imaje Er_3.SECOND" : USInt = PLC Data_DTLData."DTL_Imaje Er_3".SECOND, 1 s
   "Data_DTLData_DTL_Paper R Out[3].HOUR" : USInt = PLC Data_DTLData."DTL_Paper R Out"[3].HOUR, 1 s
   "Data_DTLData_DTL_Paper R Out[3].MINUTE" : USInt = PLC Data_DTLData."DTL_Paper R Out"[3].MINUTE, 1 s
   "Data_DTLData_DTL_Paper R Out[3].SECOND" : USInt = PLC Data_DTLData."DTL_Paper R Out"[3].SECOND, 1 s
   "Data_DTLData_DTL_Imaje Not In Position[3].HOUR" : USInt = PLC Data_DTLData."DTL_Imaje Not In Position"[3].HOUR, 1 s
   "Data_DTLData_DTL_Imaje Not In Position[3].MINUTE" : USInt = PLC Data_DTLData."DTL_Imaje Not In Position"[3].MINUTE, 1 s
   "Data_DTLData_DTL_Imaje Not In Position[3].SECOND" : USInt = PLC Data_DTLData."DTL_Imaje Not In Position"[3].SECOND, 1 s
   "DB_Integer_IDay" : USInt = PLC Data_Integer.IDay, 1 s
   "DB_Integer_IHour" : USInt = PLC Data_Integer.IHour, 1 s
   "DB_Integer_IMinute" : USInt = PLC Data_Integer.IMinute, 1 s
   "DB_Integer_IMonth" : USInt = PLC Data_Integer.IMonth, 1 s
   "DB_Integer_ISecond" : USInt = PLC Data_Integer.ISecond, 1 s
   "DB_Integer_IYear" : UInt = PLC Data_Integer.IYear, 1 s